(* Logix 5000 project; controller _GigaDiscovery vendor 1 type 14 code 244 rev 35.11; software revision 35.03; part 10 of 23 *)
(* tags used below, declared in another part *)
   Emergencies_CL1 : DINT[14];
(* S_Alarms, continued *)

ROUTINE _01_In_Out   (* ladder *)
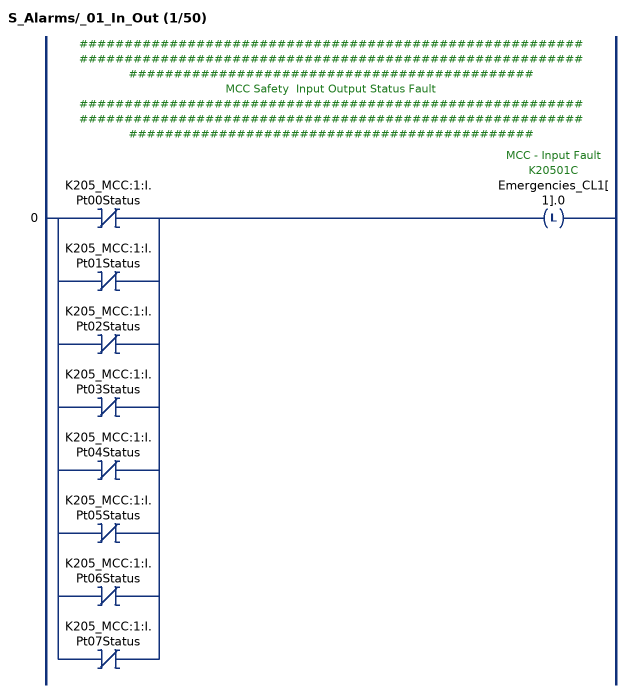
   // #############################################################################################################################################################
   // MCC Safety  Input Output Status Fault
   // #############################################################################################################################################################
   0: [XIO(K205_MCC:1:I.Pt00Status) ,XIO(K205_MCC:1:I.Pt01Status) ,XIO(K205_MCC:1:I.Pt02Status) ,XIO(K205_MCC:1:I.Pt03Status) ,XIO(K205_MCC:1:I.Pt04Status) ,XIO(K205_MCC:1:I.Pt05Status) ,XIO(K205_MCC:1:I.Pt06Status) ,XIO(K205_MCC:1:I.Pt07Status) ]OTL(Emergencies_CL1[1].0);
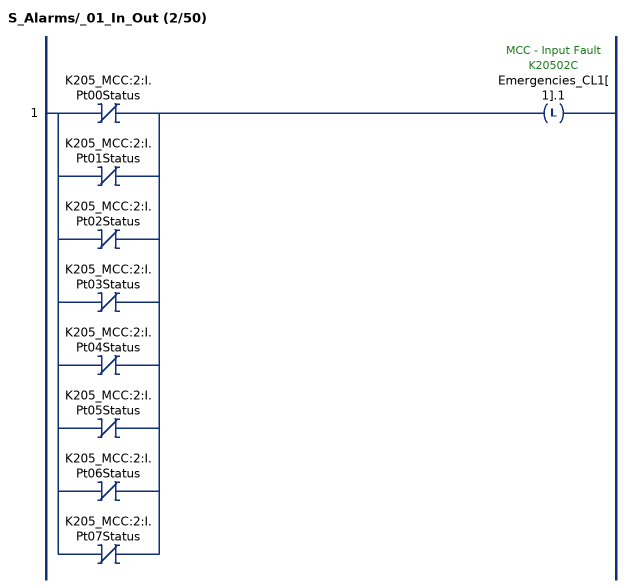
   1: [XIO(K205_MCC:2:I.Pt00Status) ,XIO(K205_MCC:2:I.Pt01Status) ,XIO(K205_MCC:2:I.Pt02Status) ,XIO(K205_MCC:2:I.Pt03Status) ,XIO(K205_MCC:2:I.Pt04Status) ,XIO(K205_MCC:2:I.Pt05Status) ,XIO(K205_MCC:2:I.Pt06Status) ,XIO(K205_MCC:2:I.Pt07Status) ]OTL(Emergencies_CL1[1].1);
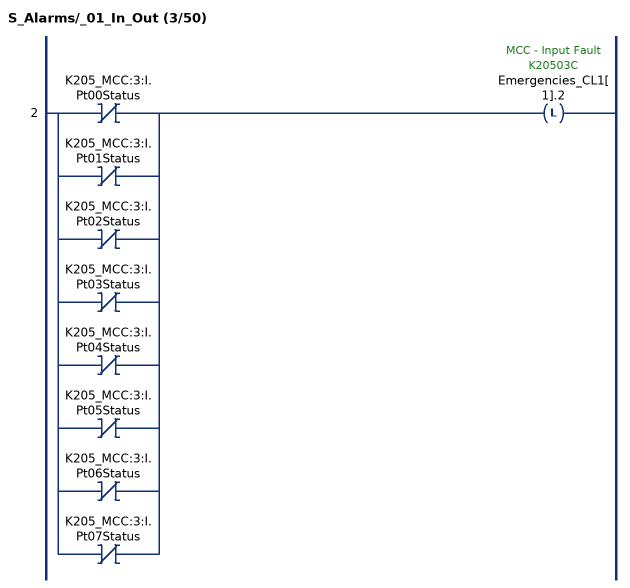
   2: [XIO(K205_MCC:3:I.Pt00Status) ,XIO(K205_MCC:3:I.Pt01Status) ,XIO(K205_MCC:3:I.Pt02Status) ,XIO(K205_MCC:3:I.Pt03Status) ,XIO(K205_MCC:3:I.Pt04Status) ,XIO(K205_MCC:3:I.Pt05Status) ,XIO(K205_MCC:3:I.Pt06Status) ,XIO(K205_MCC:3:I.Pt07Status) ]OTL(Emergencies_CL1[1].2);
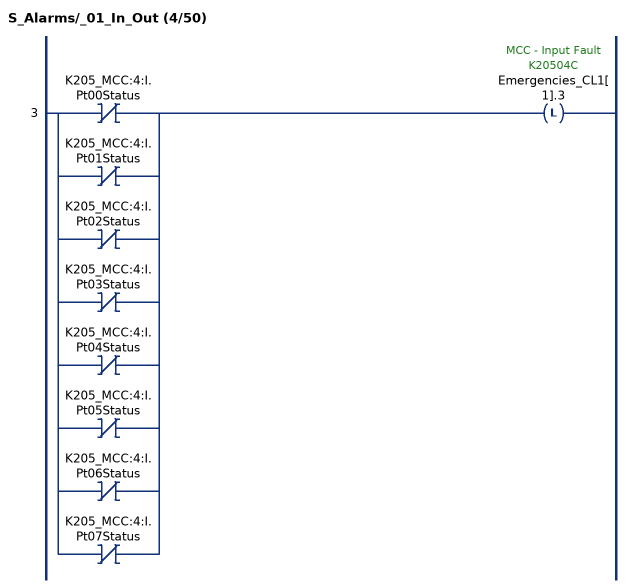
   3: [XIO(K205_MCC:4:I.Pt00Status) ,XIO(K205_MCC:4:I.Pt01Status) ,XIO(K205_MCC:4:I.Pt02Status) ,XIO(K205_MCC:4:I.Pt03Status) ,XIO(K205_MCC:4:I.Pt04Status) ,XIO(K205_MCC:4:I.Pt05Status) ,XIO(K205_MCC:4:I.Pt06Status) ,XIO(K205_MCC:4:I.Pt07Status) ]OTL(Emergencies_CL1[1].3);
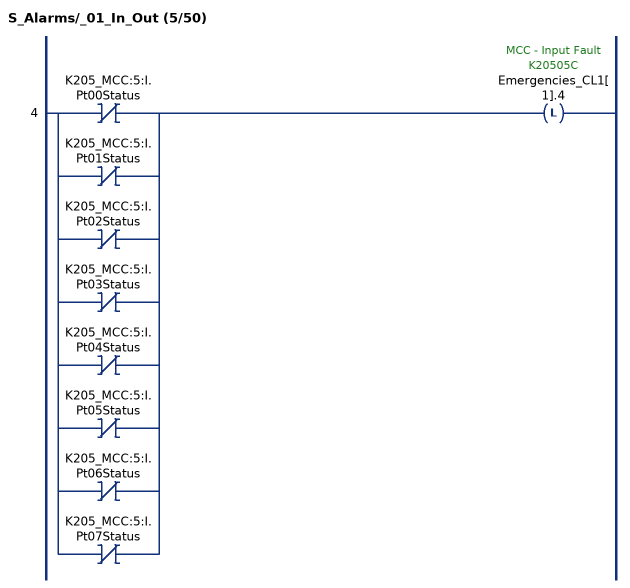
   4: [XIO(K205_MCC:5:I.Pt00Status) ,XIO(K205_MCC:5:I.Pt01Status) ,XIO(K205_MCC:5:I.Pt02Status) ,XIO(K205_MCC:5:I.Pt03Status) ,XIO(K205_MCC:5:I.Pt04Status) ,XIO(K205_MCC:5:I.Pt05Status) ,XIO(K205_MCC:5:I.Pt06Status) ,XIO(K205_MCC:5:I.Pt07Status) ]OTL(Emergencies_CL1[1].4);
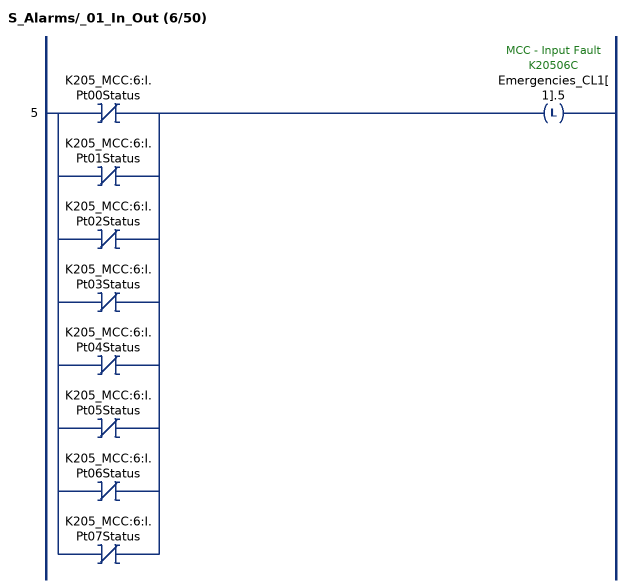
   5: [XIO(K205_MCC:6:I.Pt00Status) ,XIO(K205_MCC:6:I.Pt01Status) ,XIO(K205_MCC:6:I.Pt02Status) ,XIO(K205_MCC:6:I.Pt03Status) ,XIO(K205_MCC:6:I.Pt04Status) ,XIO(K205_MCC:6:I.Pt05Status) ,XIO(K205_MCC:6:I.Pt06Status) ,XIO(K205_MCC:6:I.Pt07Status) ]OTL(Emergencies_CL1[1].5);
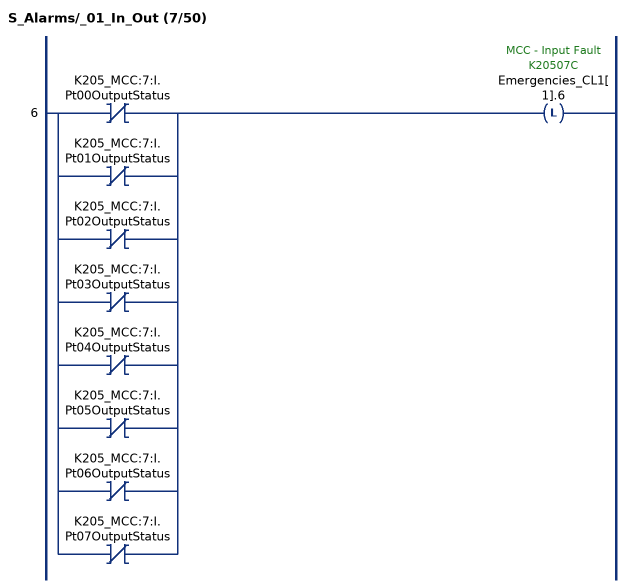
   6: [XIO(K205_MCC:7:I.Pt00OutputStatus) ,XIO(K205_MCC:7:I.Pt01OutputStatus) ,XIO(K205_MCC:7:I.Pt02OutputStatus) ,XIO(K205_MCC:7:I.Pt03OutputStatus) ,XIO(K205_MCC:7:I.Pt04OutputStatus) ,XIO(K205_MCC:7:I.Pt05OutputStatus) ,XIO(K205_MCC:7:I.Pt06OutputStatus) ,XIO(K205_MCC:7:I.Pt07OutputStatus) ]OTL(Emergencies_CL1[1].6);
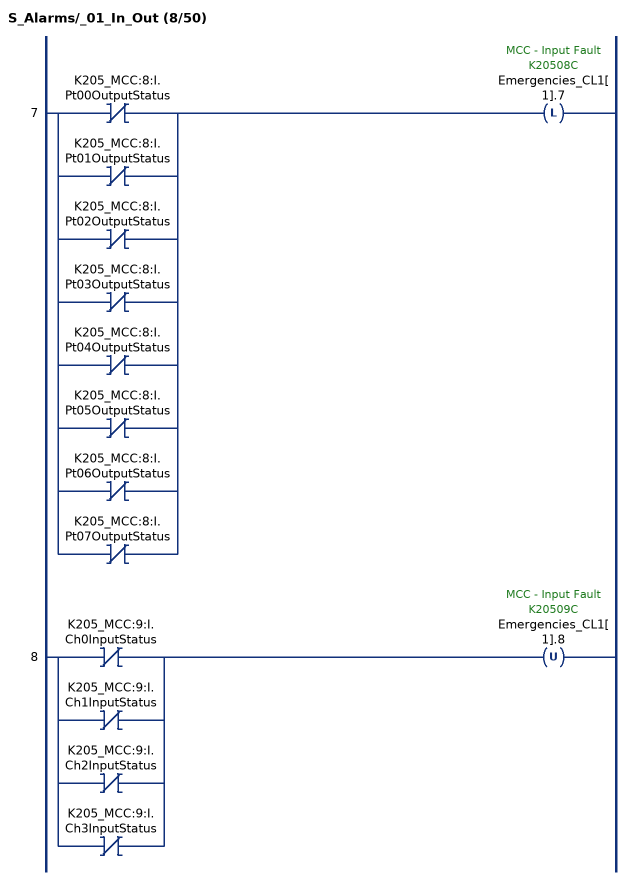
   7: [XIO(K205_MCC:8:I.Pt00OutputStatus) ,XIO(K205_MCC:8:I.Pt01OutputStatus) ,XIO(K205_MCC:8:I.Pt02OutputStatus) ,XIO(K205_MCC:8:I.Pt03OutputStatus) ,XIO(K205_MCC:8:I.Pt04OutputStatus) ,XIO(K205_MCC:8:I.Pt05OutputStatus) ,XIO(K205_MCC:8:I.Pt06OutputStatus) ,XIO(K205_MCC:8:I.Pt07OutputStatus) ]OTL(Emergencies_CL1[1].7);
   8: [XIO(K205_MCC:9:I.Ch0InputStatus) ,XIO(K205_MCC:9:I.Ch1InputStatus) ,XIO(K205_MCC:9:I.Ch2InputStatus) ,XIO(K205_MCC:9:I.Ch3InputStatus) ]OTU(Emergencies_CL1[1].8);
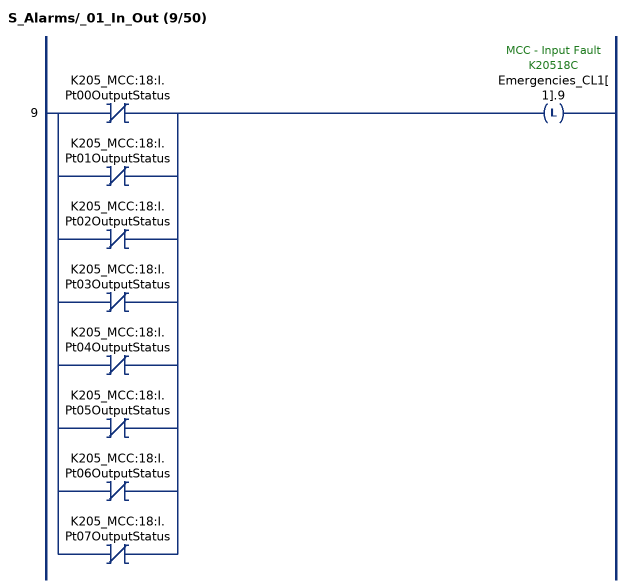
   9: [XIO(K205_MCC:18:I.Pt00OutputStatus) ,XIO(K205_MCC:18:I.Pt01OutputStatus) ,XIO(K205_MCC:18:I.Pt02OutputStatus) ,XIO(K205_MCC:18:I.Pt03OutputStatus) ,XIO(K205_MCC:18:I.Pt04OutputStatus) ,XIO(K205_MCC:18:I.Pt05OutputStatus) ,XIO(K205_MCC:18:I.Pt06OutputStatus) ,XIO(K205_MCC:18:I.Pt07OutputStatus) ]OTL(Emergencies_CL1[1].9);
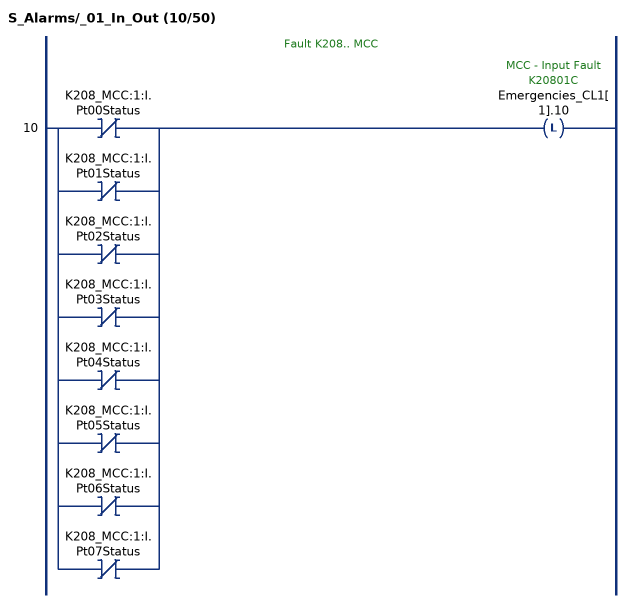
   // Fault K208.. MCC
   10: [XIO(K208_MCC:1:I.Pt00Status) ,XIO(K208_MCC:1:I.Pt01Status) ,XIO(K208_MCC:1:I.Pt02Status) ,XIO(K208_MCC:1:I.Pt03Status) ,XIO(K208_MCC:1:I.Pt04Status) ,XIO(K208_MCC:1:I.Pt05Status) ,XIO(K208_MCC:1:I.Pt06Status) ,XIO(K208_MCC:1:I.Pt07Status) ]OTL(Emergencies_CL1[1].10);
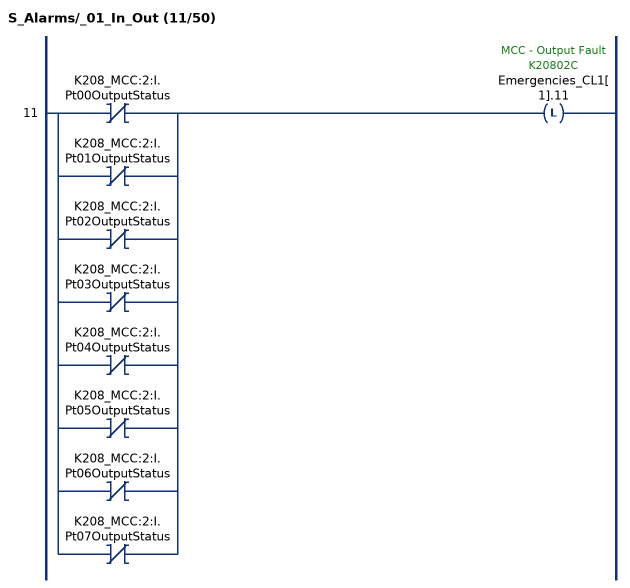
   11: [XIO(K208_MCC:2:I.Pt00OutputStatus) ,XIO(K208_MCC:2:I.Pt01OutputStatus) ,XIO(K208_MCC:2:I.Pt02OutputStatus) ,XIO(K208_MCC:2:I.Pt03OutputStatus) ,XIO(K208_MCC:2:I.Pt04OutputStatus) ,XIO(K208_MCC:2:I.Pt05OutputStatus) ,XIO(K208_MCC:2:I.Pt06OutputStatus) ,XIO(K208_MCC:2:I.Pt07OutputStatus) ]OTL(Emergencies_CL1[1].11);
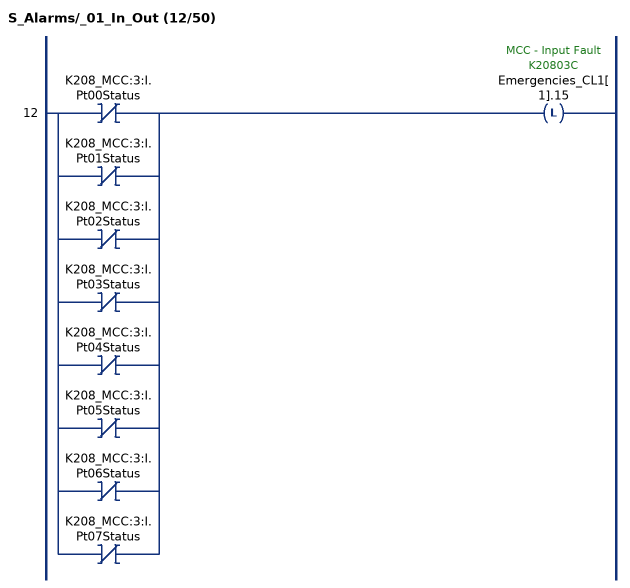
   12: [XIO(K208_MCC:3:I.Pt00Status) ,XIO(K208_MCC:3:I.Pt01Status) ,XIO(K208_MCC:3:I.Pt02Status) ,XIO(K208_MCC:3:I.Pt03Status) ,XIO(K208_MCC:3:I.Pt04Status) ,XIO(K208_MCC:3:I.Pt05Status) ,XIO(K208_MCC:3:I.Pt06Status) ,XIO(K208_MCC:3:I.Pt07Status) ]OTL(Emergencies_CL1[1].15);
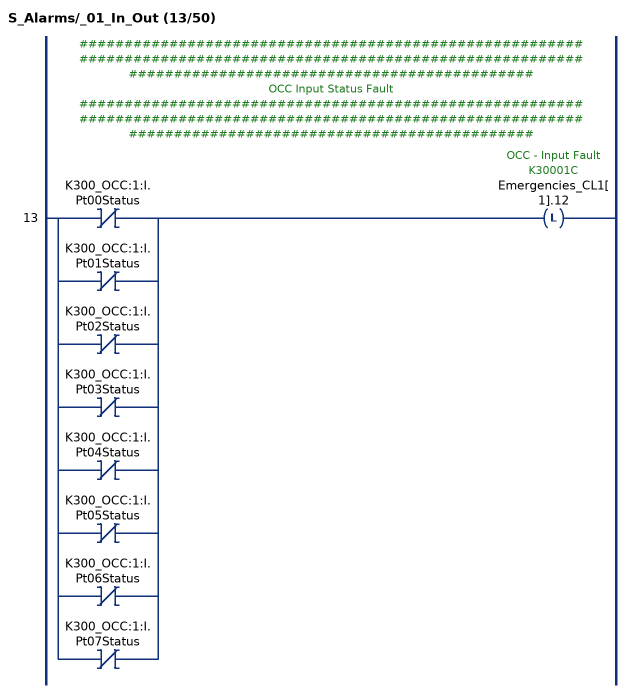
   // #############################################################################################################################################################
   // OCC Input Status Fault
   // #############################################################################################################################################################
   13: [XIO(K300_OCC:1:I.Pt00Status) ,XIO(K300_OCC:1:I.Pt01Status) ,XIO(K300_OCC:1:I.Pt02Status) ,XIO(K300_OCC:1:I.Pt03Status) ,XIO(K300_OCC:1:I.Pt04Status) ,XIO(K300_OCC:1:I.Pt05Status) ,XIO(K300_OCC:1:I.Pt06Status) ,XIO(K300_OCC:1:I.Pt07Status) ]OTL(Emergencies_CL1[1].12);
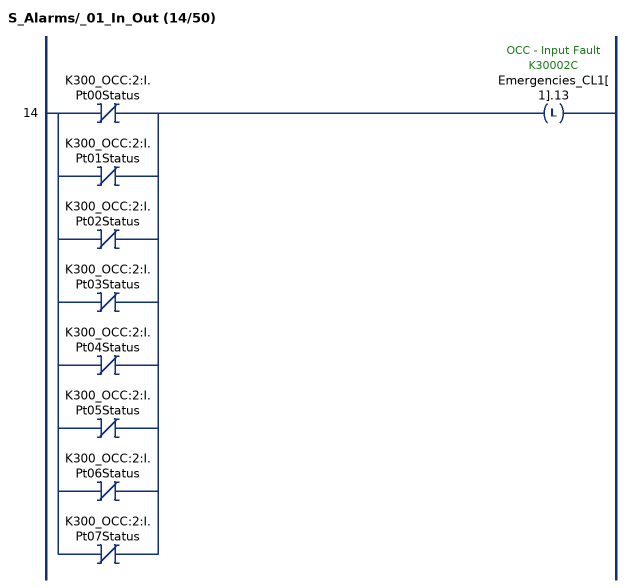
   14: [XIO(K300_OCC:2:I.Pt00Status) ,XIO(K300_OCC:2:I.Pt01Status) ,XIO(K300_OCC:2:I.Pt02Status) ,XIO(K300_OCC:2:I.Pt03Status) ,XIO(K300_OCC:2:I.Pt04Status) ,XIO(K300_OCC:2:I.Pt05Status) ,XIO(K300_OCC:2:I.Pt06Status) ,XIO(K300_OCC:2:I.Pt07Status) ]OTL(Emergencies_CL1[1].13);
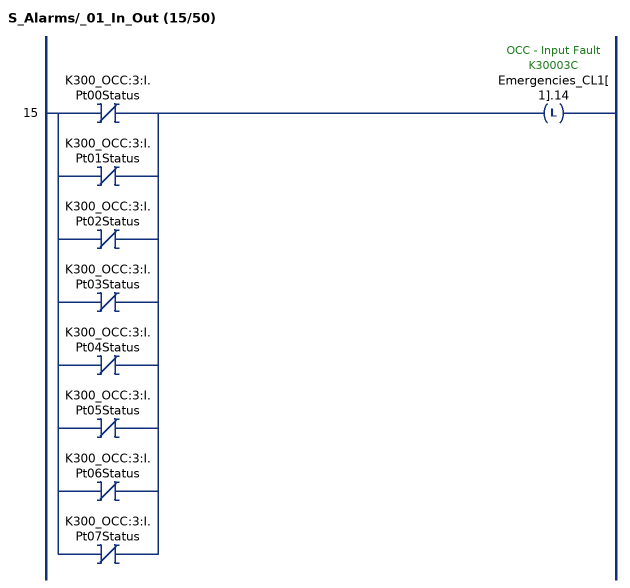
   15: [XIO(K300_OCC:3:I.Pt00Status) ,XIO(K300_OCC:3:I.Pt01Status) ,XIO(K300_OCC:3:I.Pt02Status) ,XIO(K300_OCC:3:I.Pt03Status) ,XIO(K300_OCC:3:I.Pt04Status) ,XIO(K300_OCC:3:I.Pt05Status) ,XIO(K300_OCC:3:I.Pt06Status) ,XIO(K300_OCC:3:I.Pt07Status) ]OTL(Emergencies_CL1[1].14);
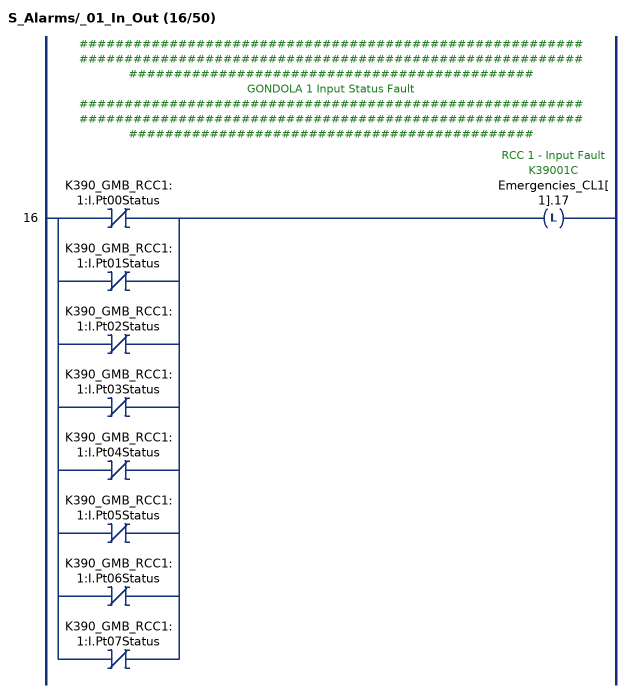
   // #############################################################################################################################################################
   // GONDOLA 1 Input Status Fault
   // #############################################################################################################################################################
   16: [XIO(K390_GMB_RCC1:1:I.Pt00Status) ,XIO(K390_GMB_RCC1:1:I.Pt01Status) ,XIO(K390_GMB_RCC1:1:I.Pt02Status) ,XIO(K390_GMB_RCC1:1:I.Pt03Status) ,XIO(K390_GMB_RCC1:1:I.Pt04Status) ,XIO(K390_GMB_RCC1:1:I.Pt05Status) ,XIO(K390_GMB_RCC1:1:I.Pt06Status) ,XIO(K390_GMB_RCC1:1:I.Pt07Status) ]OTL(Emergencies_CL1[1].17);
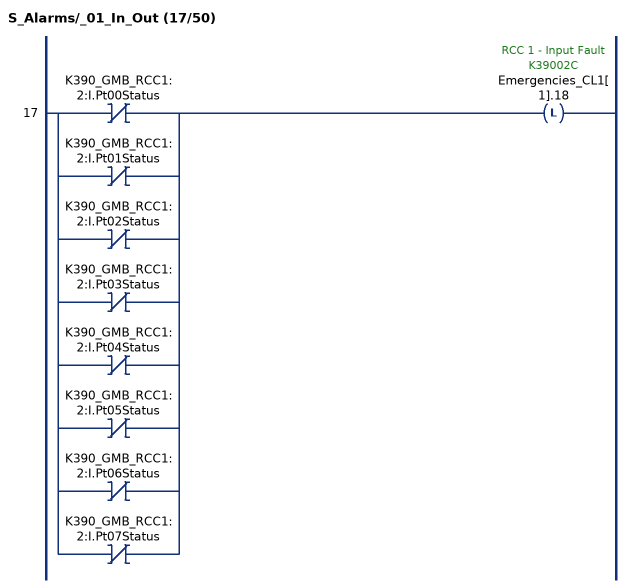
   17: [XIO(K390_GMB_RCC1:2:I.Pt00Status) ,XIO(K390_GMB_RCC1:2:I.Pt01Status) ,XIO(K390_GMB_RCC1:2:I.Pt02Status) ,XIO(K390_GMB_RCC1:2:I.Pt03Status) ,XIO(K390_GMB_RCC1:2:I.Pt04Status) ,XIO(K390_GMB_RCC1:2:I.Pt05Status) ,XIO(K390_GMB_RCC1:2:I.Pt06Status) ,XIO(K390_GMB_RCC1:2:I.Pt07Status) ]OTL(Emergencies_CL1[1].18);
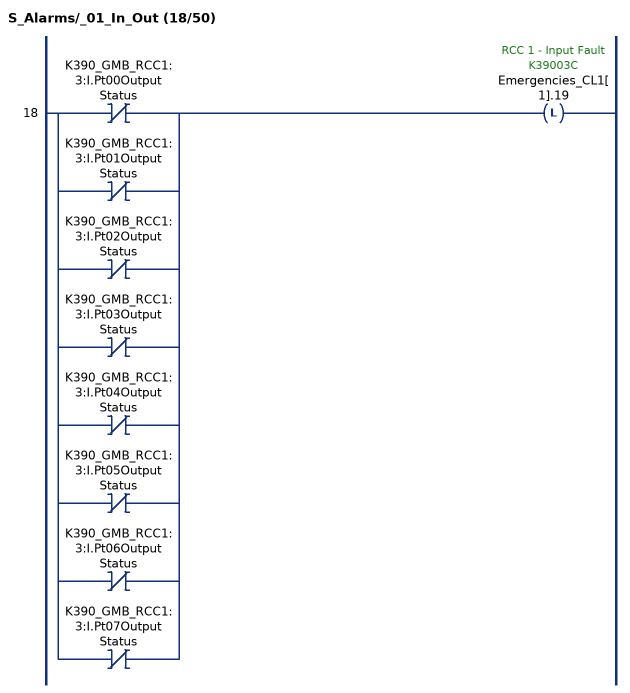
   18: [XIO(K390_GMB_RCC1:3:I.Pt00OutputStatus) ,XIO(K390_GMB_RCC1:3:I.Pt01OutputStatus) ,XIO(K390_GMB_RCC1:3:I.Pt02OutputStatus) ,XIO(K390_GMB_RCC1:3:I.Pt03OutputStatus) ,XIO(K390_GMB_RCC1:3:I.Pt04OutputStatus) ,XIO(K390_GMB_RCC1:3:I.Pt05OutputStatus) ,XIO(K390_GMB_RCC1:3:I.Pt06OutputStatus) ,XIO(K390_GMB_RCC1:3:I.Pt07OutputStatus) ]OTL(Emergencies_CL1[1].19);
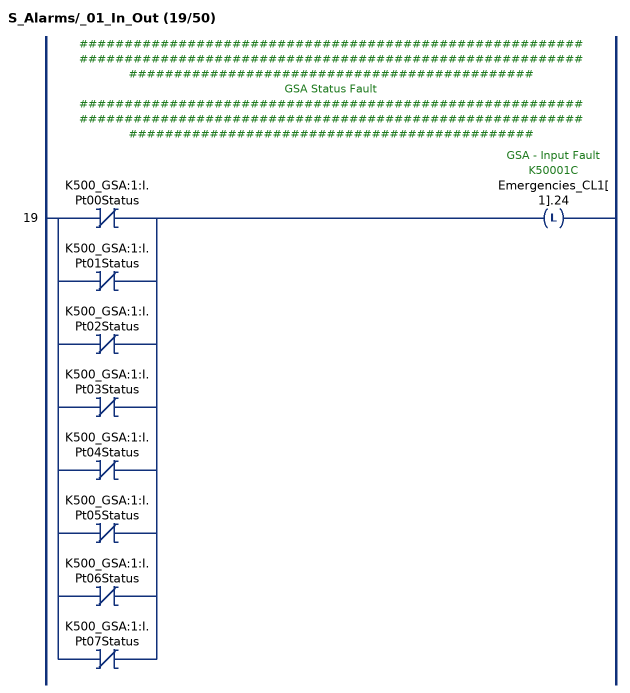
   // #############################################################################################################################################################
   // GSA Status Fault
   // #############################################################################################################################################################
   19: [XIO(K500_GSA:1:I.Pt00Status) ,XIO(K500_GSA:1:I.Pt01Status) ,XIO(K500_GSA:1:I.Pt02Status) ,XIO(K500_GSA:1:I.Pt03Status) ,XIO(K500_GSA:1:I.Pt04Status) ,XIO(K500_GSA:1:I.Pt05Status) ,XIO(K500_GSA:1:I.Pt06Status) ,XIO(K500_GSA:1:I.Pt07Status) ]OTL(Emergencies_CL1[1].24);
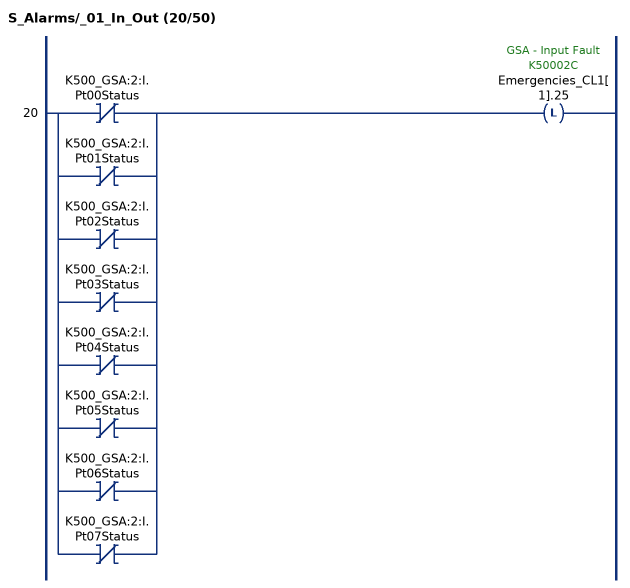
   20: [XIO(K500_GSA:2:I.Pt00Status) ,XIO(K500_GSA:2:I.Pt01Status) ,XIO(K500_GSA:2:I.Pt02Status) ,XIO(K500_GSA:2:I.Pt03Status) ,XIO(K500_GSA:2:I.Pt04Status) ,XIO(K500_GSA:2:I.Pt05Status) ,XIO(K500_GSA:2:I.Pt06Status) ,XIO(K500_GSA:2:I.Pt07Status) ]OTL(Emergencies_CL1[1].25);
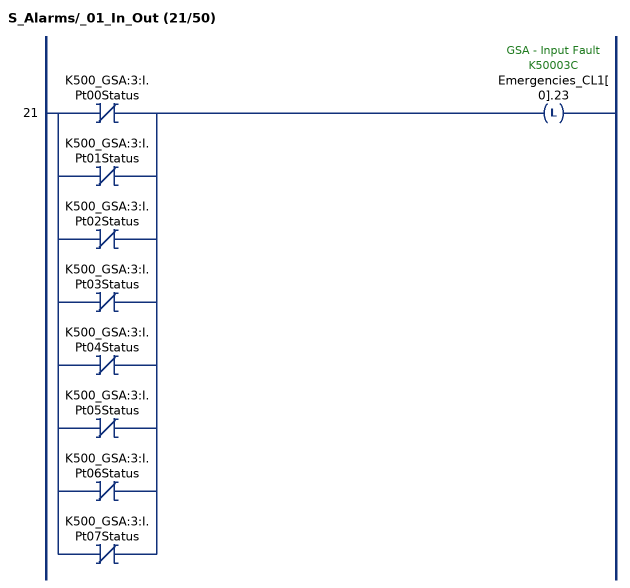
   21: [XIO(K500_GSA:3:I.Pt00Status) ,XIO(K500_GSA:3:I.Pt01Status) ,XIO(K500_GSA:3:I.Pt02Status) ,XIO(K500_GSA:3:I.Pt03Status) ,XIO(K500_GSA:3:I.Pt04Status) ,XIO(K500_GSA:3:I.Pt05Status) ,XIO(K500_GSA:3:I.Pt06Status) ,XIO(K500_GSA:3:I.Pt07Status) ]OTL(Emergencies_CL1[0].23);
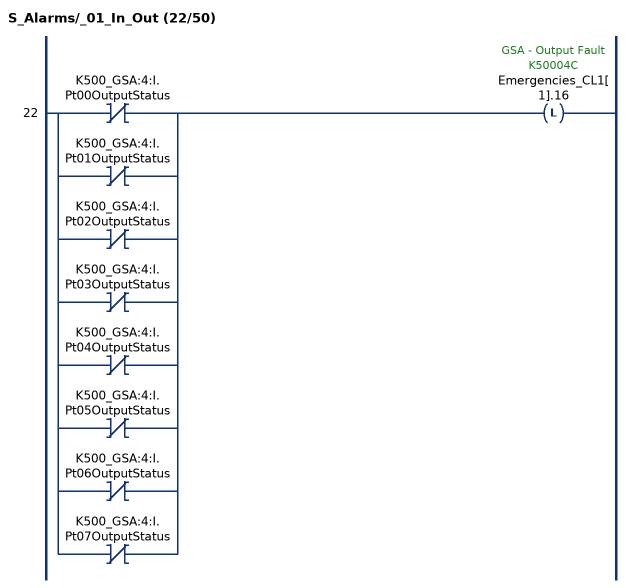
   22: [XIO(K500_GSA:4:I.Pt00OutputStatus) ,XIO(K500_GSA:4:I.Pt01OutputStatus) ,XIO(K500_GSA:4:I.Pt02OutputStatus) ,XIO(K500_GSA:4:I.Pt03OutputStatus) ,XIO(K500_GSA:4:I.Pt04OutputStatus) ,XIO(K500_GSA:4:I.Pt05OutputStatus) ,XIO(K500_GSA:4:I.Pt06OutputStatus) ,XIO(K500_GSA:4:I.Pt07OutputStatus) ]OTL(Emergencies_CL1[1].16);
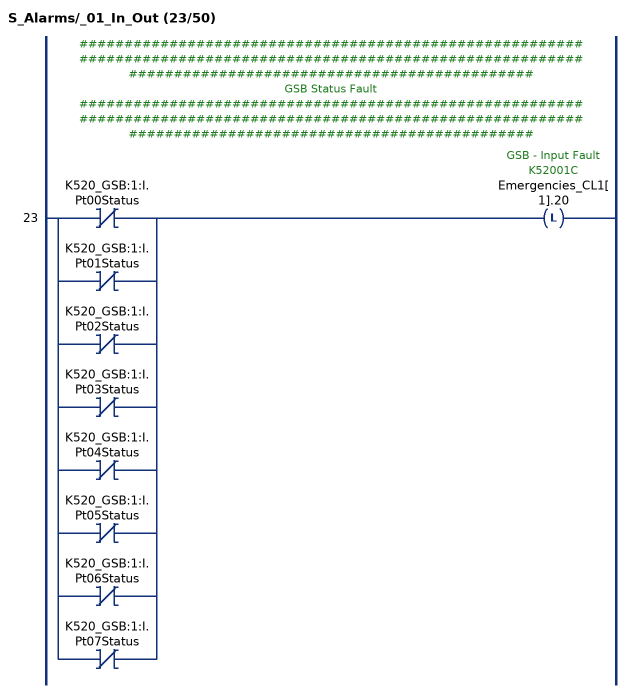
   // #############################################################################################################################################################
   // GSB Status Fault
   // #############################################################################################################################################################
   23: [XIO(K520_GSB:1:I.Pt00Status) ,XIO(K520_GSB:1:I.Pt01Status) ,XIO(K520_GSB:1:I.Pt02Status) ,XIO(K520_GSB:1:I.Pt03Status) ,XIO(K520_GSB:1:I.Pt04Status) ,XIO(K520_GSB:1:I.Pt05Status) ,XIO(K520_GSB:1:I.Pt06Status) ,XIO(K520_GSB:1:I.Pt07Status) ]OTL(Emergencies_CL1[1].20);
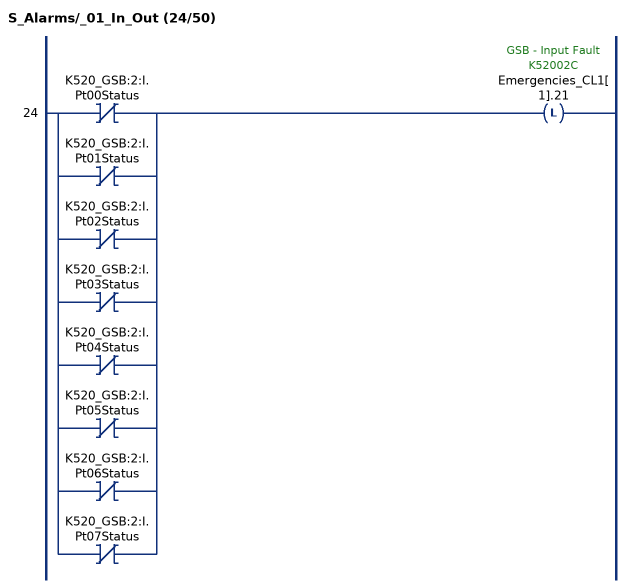
   24: [XIO(K520_GSB:2:I.Pt00Status) ,XIO(K520_GSB:2:I.Pt01Status) ,XIO(K520_GSB:2:I.Pt02Status) ,XIO(K520_GSB:2:I.Pt03Status) ,XIO(K520_GSB:2:I.Pt04Status) ,XIO(K520_GSB:2:I.Pt05Status) ,XIO(K520_GSB:2:I.Pt06Status) ,XIO(K520_GSB:2:I.Pt07Status) ]OTL(Emergencies_CL1[1].21);
